// TIA Portal project "1215C_BREAKOUT_BOARD_IO-LINK_TOWERLIGHT" (V19) (continued)
REGION Network 6: Saving Selections
   RUNG wire#powerrail
      Contact( "DB005-HMI_Data".TowerLight.xSave_Config )
      wire#w1
      Move(in := #Seg2.iTempAnimation, out1 => "DB005-HMI_Data".TowerLight.Segment2.iSavedAnimate)
      Move(in := #Seg2.iTempSpeed, out1 => "DB003-IOLink_I/O".Outputs.TL_Byte_Array[13])
   END_RUNG
   RUNG wire#w1
      Move(in := #Seg2.iTempColour1, out1 => "DB003-IOLink_I/O".Outputs.TL_Byte_Array[15])
      Move(in := #Seg2.iTempColour2, out1 => "DB003-IOLink_I/O".Outputs.TL_Byte_Array[14])
      Move(in := #Seg2."iTempClrWidth%", out1 => "DB003-IOLink_I/O".Outputs.TL_Byte_Array[12])
   END_RUNG
   // the same network as SCL:
   IF "DB005-HMI_Data".TowerLight.xSave_Config THEN
       "DB005-HMI_Data".TowerLight.Segment2.iSavedAnimate := #Seg2.iTempAnimation;
       "DB003-IOLink_I/O".Outputs.TL_Byte_Array[13] := #Seg2.iTempSpeed;
       "DB003-IOLink_I/O".Outputs.TL_Byte_Array[15] := #Seg2.iTempColour1;
       "DB003-IOLink_I/O".Outputs.TL_Byte_Array[14] := #Seg2.iTempColour2;
       "DB003-IOLink_I/O".Outputs.TL_Byte_Array[12] := #Seg2."iTempClrWidth%";
   END_IF;
END_REGION

REGION Network 7: ================= SEGMENT_THREE =================
END_REGION

REGION Network 8: While making selections
   RUNG wire#powerrail
      { S7_Templates := "SrcType := UInt" } EQ_Contact(in1 := "DB005-HMI_Data".iScreen_Number, in2 := 9)
      wire#w1
      Move(in := "DB005-HMI_Data".TowerLight.Segment3.iAnimate, out1 => #Seg3.iTempAnimation)
      Move(in := "DB005-HMI_Data".TowerLight.Segment3.iSpeed, out1 => #Seg3.iTempSpeed)
   END_RUNG
   RUNG wire#w1
      Move(in := "DB005-HMI_Data".TowerLight.Segment3.iColour1, out1 => #Seg3.iTempColour1)
      Move(in := "DB005-HMI_Data".TowerLight.Segment3.iColour2, out1 => #Seg3.iTempColour2)
      Move(in := "DB005-HMI_Data".TowerLight.Segment3."iClrWidth%", out1 => #Seg3."iTempClrWidth%")
   END_RUNG
   // the same network as SCL:
   IF "DB005-HMI_Data".iScreen_Number = 9 THEN
       #Seg3.iTempAnimation := "DB005-HMI_Data".TowerLight.Segment3.iAnimate;
       #Seg3.iTempSpeed := "DB005-HMI_Data".TowerLight.Segment3.iSpeed;
       #Seg3.iTempColour1 := "DB005-HMI_Data".TowerLight.Segment3.iColour1;
       #Seg3.iTempColour2 := "DB005-HMI_Data".TowerLight.Segment3.iColour2;
       #Seg3."iTempClrWidth%" := "DB005-HMI_Data".TowerLight.Segment3."iClrWidth%";
   END_IF;
END_REGION

REGION Network 9: Saving Selections
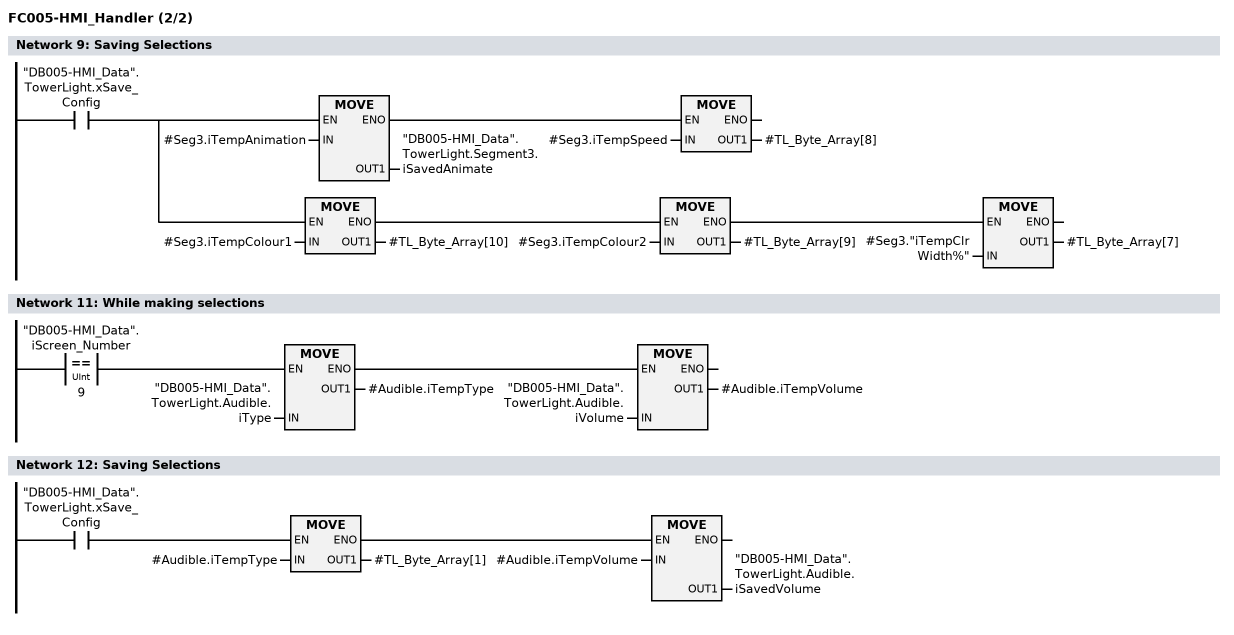
   RUNG wire#powerrail
      Contact( "DB005-HMI_Data".TowerLight.xSave_Config )
      wire#w1
      Move(in := #Seg3.iTempAnimation, out1 => "DB005-HMI_Data".TowerLight.Segment3.iSavedAnimate)
      Move(in := #Seg3.iTempSpeed, out1 => #TL_Byte_Array[8])
   END_RUNG
   RUNG wire#w1
      Move(in := #Seg3.iTempColour1, out1 => #TL_Byte_Array[10])
      Move(in := #Seg3.iTempColour2, out1 => #TL_Byte_Array[9])
      Move(in := #Seg3."iTempClrWidth%", out1 => #TL_Byte_Array[7])
   END_RUNG
   // the same network as SCL:
   IF "DB005-HMI_Data".TowerLight.xSave_Config THEN
       "DB005-HMI_Data".TowerLight.Segment3.iSavedAnimate := #Seg3.iTempAnimation;
       #TL_Byte_Array[8] := #Seg3.iTempSpeed;
       #TL_Byte_Array[10] := #Seg3.iTempColour1;
       #TL_Byte_Array[9] := #Seg3.iTempColour2;
       #TL_Byte_Array[7] := #Seg3."iTempClrWidth%";
   END_IF;
END_REGION

REGION Network 10: ================= AUDIBLE =================
END_REGION

REGION Network 11: While making selections
   RUNG wire#powerrail
      { S7_Templates := "SrcType := UInt" } EQ_Contact(in1 := "DB005-HMI_Data".iScreen_Number, in2 := 9)
      Move(in := "DB005-HMI_Data".TowerLight.Audible.iType, out1 => #Audible.iTempType)
      Move(in := "DB005-HMI_Data".TowerLight.Audible.iVolume, out1 => #Audible.iTempVolume)
   END_RUNG
   // the same network as SCL:
   IF "DB005-HMI_Data".iScreen_Number = 9 THEN
       #Audible.iTempType := "DB005-HMI_Data".TowerLight.Audible.iType;
       #Audible.iTempVolume := "DB005-HMI_Data".TowerLight.Audible.iVolume;
   END_IF;
END_REGION

REGION Network 12: Saving Selections
   RUNG wire#powerrail
      Contact( "DB005-HMI_Data".TowerLight.xSave_Config )
      Move(in := #Audible.iTempType, out1 => #TL_Byte_Array[1])
      Move(in := #Audible.iTempVolume, out1 => "DB005-HMI_Data".TowerLight.Audible.iSavedVolume)
   END_RUNG
   // the same network as SCL:
   IF "DB005-HMI_Data".TowerLight.xSave_Config THEN
       #TL_Byte_Array[1] := #Audible.iTempType;
       "DB005-HMI_Data".TowerLight.Audible.iSavedVolume := #Audible.iTempVolume;
   END_IF;
END_REGION
END_FUNCTION

// ===== library types =====

// folder: S7-1200/1500/Lib/S7-1200/1500/Common

FUNCTION_BLOCK "IO_LINK_DEVICE"   // FB50001, SCL
TITLE = IO_LINK_DEVICE
{ S7_Optimized_Access := 'TRUE' }
AUTHOR : SUP_FA
FAMILY : IO-Link
VERSION : 3.0
// Function block to read and write acyclic data on devices with IO-Link used on SIMATIC S7 controllers. (former IO_LINK_CALL)
   VAR_INPUT
      REQ : Bool;   // request function / Request Function / Neuer Auftrag
      ID : HW_IO;   // hardware identifier of IO-Link master module (HW_IO) from hw-config / Hardwarekennung des IOL-Master Moduls (HW_IO) aus HW-Konfiguration
      CAP : DInt := DINT#0;   // Client Access Point (CAP), for ET200 always 227 decimal / Client Access Point (CAP), bei ET200 immer 227 dez
      RD_WR : Bool;   // read and write access on IO-Link device 0: read, 1: write / Lese und Schreibzugriff auf IO-Link Device 0: Lesen, 1: schreiben
      PORT : Int := INT#0;   // number of port on IO-Link master module (ET200SP = 0..4) / Port/ Kanalnummer an dem das IO-Link Device betrieben wird. (ET200 = 0 .. 4)
      IOL_INDEX : Int := INT#0;   // address parameter Index (IO-Link Device) 0..32767 IOL-D, 65535 port functions / Adressparameter Index (IO-Link Device) 0..32767 IOL-D, 65535 port functions
      IOL_SUBINDEX : Int := INT#0;   // address parameter Subindex (IO-Link Device) 0 full record; 1-255 single parameter / Adressparameter Subindex (IO-Link Device) 0 ges. Record; 1-255 einz. Parameter
      LEN : Int := INT#0;   // length of writing data (netto data) / Länge der zu schreibenden Daten (Nettodaten)
   END_VAR
   VAR_OUTPUT
      DONE_VALID : Bool;   // validity 0: data invalid ; 1: data valid / Gültigkeit 0: Daten nicht gültig; 1: Daten gültig
      BUSY : Bool;   // 0: request finish 1: request in progress / 0: Auftrag abgeschlossen 1: Auftrag in Bearbeitung
      ERROR : Bool;   // Error Flag = 0: no error; 1: function aborted with error / Fehler Flag 0: kein Fehler; 1: Abbruch der Funktion mit Fehler
      STATUS : DWord := DW#16#00000000;   // DP/ PNIO - error status ; ERROR Flag = 1 - communication error status in detail / DP/ PNIO - Fehlerstatus; ERROR Flag = 1 - detaillierter Kommunikationsfehlerstatus
      IOL_STATUS : DWord := DW#16#00000000;   // IO-Link error status; ERROR flag = 1: IO-Link error status in detail / IO-Link Fehlerstatus; ERROR Flag = 1 - detaillierte IO-Link Fehlerstatus
      RD_LEN : Int := INT#0;   // length of read data record (number of bytes) / Länge des gelesenen Datensatzes (Anzahl Bytes)
   END_VAR
   VAR_IN_OUT
      RECORD_IOL_DATA : Array[0..231] of Byte;   // data area for reading / writing data (max. 232 byte) / Datenbereich für LESEN / SCHREIBEN (max. 232 Byte)
   END_VAR
   VAR
      RDREC_Function : RDREC;   // system function "read data record" (former SFB52) / Funktion Datensatz lesen (ehemals SFB52)
      WRREC_Function : WRREC;   // system function "write data record" (former SFB53) / Funktion Datensatz schreiben (ehemals SFB53)
      TP_poll : TP_TIME;   // poll rate read data record / Pollzeit für "Datensatz lesen"
      TON_monitoring : TON_TIME;   // request monitoring time / Überwachungszeit für Aufträge
      rdrec : Struct   // internal structure for RDREC / interne Struktur für RDREC
         valid : Bool;   // Function performed
         busy : Bool;   // Function busy
         error : Bool;   // Error flag
         status : DWord;   // Function result/error message
         length : UInt;   // Length of the fetched data record
      END_STRUCT;
      wrrec : Struct   // internal structure for WRREC / interne Struktur für WRREC
         length : UInt;   // length of write data record
         done : Bool;   // Function performed
         busy : Bool;   // Function busy
         error : Bool;   // Error flag
         status : DWord;   // Function result/error message
      END_STRUCT;
      read : Struct   // data area for reading data / Datenbereich für Lesedaten
         header : Struct
            CALL : Struct   // header for read/write data record
               Extended_Function_Num : Byte := 16#8;   // extended function number (fix coded 08h)
               Port : Byte;   // variable port (user interface) 0...255
               FI_Index : Word := 16#FE4A;   // FI index (fix coded 65098)
            END_STRUCT;
            IOL : Struct   // header for IO-Link
               Control : Byte;   // RD_WR = 0 = read = Control:=0x03 / / RD_WR = 1 = write = Control:=0x02
               Index_HighByte : Byte;   // index of data record 0…32767 (high byte)
               Index_LowByte : Byte;   // index of data record 0…32767 (low byte)
               Subindex : Byte;   // subindex for data record 0...255
            END_STRUCT;
         END_STRUCT;
         data : Array[0..231] of Byte;
      END_STRUCT;
      write : Struct   // data area for writing data / Datenbereich für Schreibdaten
         header : Struct
            CALL : Struct   // header for read/write data record
               Extended_Function_Num : Byte := 16#8;   // extended function number (fix coded 08h)
               Port : Byte;   // variable port (user interface) 0...255
               FI_Index : Word := 16#FE4A;   // FI index (fix coded 65098)
            END_STRUCT;
            IOL : Struct   // header for IO-Link
               Control : Byte;   // RD_WR = 0 = read = Control:=0x03 / / RD_WR = 1 = write = Control:=0x02
               Index_HighByte : Byte;   // index of data record 0…32767 (high byte)
               Index_LowByte : Byte;   // index of data record 0…32767 (low byte)
               Subindex : Byte;   // subindex for data record 0...255
            END_STRUCT;
         END_STRUCT;
         data : Array[0..231] of Byte;
      END_STRUCT;
      sequencecontrol : Int := INT#0;   // number of sequence control
      typeofrequest : Int := INT#0;   // type of request (0=Read, 1=Write)
      R_TRIG_REQ : Bool;   // impulse start new request / Impuls für neuen Auftrag starten
      R_TRIG_REQ_old : Bool;   // old value of REQ (previous cycle) / Flankenmerker
      F_TRIG_poll : Bool;   // impulse poll read data record (response) / Impuls für Pollen "Datensatz lesen"
      F_TRIG_poll_old : Bool;   // old value of Poll (previous cycle) / Flankenmerker
   END_VAR
   VAR_TEMP
      retval : Int;   // function return value / Variable für Rückgabewerte von Funktionen
      tmpWORD : Word;   // data type WORD for temporarily use / Datentyp WORD zur temporären Verwendung
      tmpDWORD : DWord;   // data type DWORD for temporarily use / Datentyp DWORD zur temporären Verwendung
      tmpINT : Int;   // data type INT for temporarily use / Datentyp INT zur temporären Verwendung
      i : Int;   // run tag for counting loops / Laufvariable für for-Schleifen
   END_VAR
BEGIN
   (*---------------------------------------------------------------------------------------------------------------------
   SIEMENS AG
   ©Copyright 2015. All Rights Reserved.
   -----------------------------------------------------------------------------------------------------------------------
   Limitation of liability
   This software was developed with largest care. However, the author can not guarantee, that the software runs under
   each version of STEP7 on each PLC flawlessly.
   There is no warranty for the software, to the extent permitted by applicable law. The copyright holder provides the
   software "as is" without warranty of any kind, either expressed or implied, including, but not limited to, the implied
   warranties of merchantability and fitness for a particular purpose. The entire risk as to the quality and performance
   of the software is with you. Should the software prove defective, you assume the cost of all necessary servicing,
   repair or correction. In no event unless required by applicable law will the copyright holder be liable to you for
   damages, including any general, special, incidental or consequential damages arising out of the use or inability to
   use the software (including but not limited to loss of data or data being rendered inaccurate or losses sustained by
   you or third parties or a failure of the software to operate with any other programs), even if such holder or other
   party has been advised of the possibility of such damages.
   Permission to use or copy this software for any purpose is hereby granted without fee, provided the above notices are
   retained on all copies. Permission to modify the code and to distribute modified code is granted, provided the above
   notices are retained, and a notice that the code was modified is included with the above copyright notice.
   -----------------------------------------------------------------------------------------------------------------------
   Functionality provided by this source (short description):
   Function block IO_LINK_DEVICE - used to read and write of acyclic data records on devices with IO-Link.
   Note:
   To read data records, the IO-Link master modules needs to know which data record is required. Therefore it is necessary
   to send at first a request via write data record (only header of 8 byte). As response the IO-Link master module
   will send the required data record.

   Status:     Released (tested)
   File name:  IO_LINK_DEVICE
   System :    SIMATIC S7-1200/1500
   Version :   3.0
   -----------------------------------------------------------------------------------------------------------------------
   Script to be stored on level ... in project (mark appropriate levels with [x] below)
   [ ] External
   [ ] All levels possible
   [x] Project level
   [ ] Controller level
   [ ] Device level
   [ ] Subobject level
   -----------------------------------------------------------------------------------------------------------------------
   Restrictions, known limitations:
   The limitation of 240 byte is based on PROFIBUS DP protocol. With PROFINET IO there wouldn't no limit but because of 
   compatibility reason it wasn't changed.
     - header =   8 byte
     - data   = 232 byte
   -----------------------------------------------------------------------------------------------------------------------
   Requirements, prerequisites, External resources used: nothing
   -----------------------------------------------------------------------------------------------------------------------
   Change log table (latest change is at the bottom OF the list):
   Version Date Changes applied
   V2.0.0 <2013-09-30> First created with TIA Portal V12 SP1
   V2.1.0 <2014-03-14> Upgrade system function 'WRREC' from V1.0 to V1.1 and released for TIA Portal V13
   V3.0.0 <2015-02-28> Upgrade and released for TIA Portal V13 SP1 (without backup/restore master parameter)
   V3.0.2 <2015-07-07> Change of #IOL_INDEX and #Port lower boundry to 0
   ---------------------------------------------------------------------------------------------------------------------*)

   (*---------------------------------------------------------------------------------------------------------------------
   Description of programmed IO-Link error codes
   8000 = time out
   8001 = wrong port
   8002 = wrong index
   8003 = wrong subindex
   8005 = wrong length for write data record
   8006 = wrong length for read data record
   8052 = error during reading data record
   8053 = error during writing data record
   All other codes are coming from a higher level!
   ---------------------------------------------------------------------------------------------------------------------*)

   (*---------------------------------------------------------------------------------------------------------------------
               NEW REQUEST
   ---------------------------------------------------------------------------------------------------------------------*)
   // detection rising edge of "REQ"
   #R_TRIG_REQ := #REQ = TRUE AND #R_TRIG_REQ_old = FALSE;
   #R_TRIG_REQ_old := #REQ = TRUE;

   // start new request if not busy
   IF #R_TRIG_REQ = TRUE AND #sequencecontrol = 0 THEN
       // Freeze record ID and CAP
       #WRREC_Function.ID := #ID;
       #WRREC_Function.INDEX := #CAP;
       #RDREC_Function.ID := #ID;
       #RDREC_Function.INDEX := #CAP;

       // Initialize outputs
       #DONE_VALID := FALSE;
       #BUSY := TRUE;
       #ERROR := FALSE;
       #STATUS := DW#16#00000000;
       #IOL_STATUS := DW#16#00000000;
       #RD_LEN := INT#0;

       // Initialize data area
       #read.header.CALL.Port := B#16#0;
       #read.header.IOL.Index_LowByte := B#16#0;
       #read.header.IOL.Index_HighByte := B#16#0;
       #read.header.IOL.Subindex := B#16#0;
       #i := INT#0; // initialize loop counter      
       FOR #i := 0 TO 231 DO
           #write.data[#i] := B#16#0;
           #read.data[#i] := B#16#0;
       END_FOR;

   (*---------------------------------------------------------------------------------------------------------------------
       Setup IO-LINK Call needs a specific header
   ---------------------------------------------------------------------------------------------------------------------*)
   // setup CALL header
   #write.header.CALL.Extended_Function_Num := 16#08;  // extended function number (fix coded 08h)
   #write.header.CALL.Port := INT_TO_BYTE(#PORT);  // 1..63 = PORT number, 64..255=reserved
   #write.header.CALL.FI_Index := 65098;  // IOL-Header is following (fix coded 65098)

   // setup IOL header 
   // CONTROL = please see below at BODY
   // INDEX
   #write.header.IOL.Index_LowByte := INT_TO_BYTE(#IOL_INDEX);
   #tmpWORD := INT_TO_WORD(#IOL_INDEX);
   #tmpWORD := SHR(IN := #tmpWORD, N := 8);
   #write.header.IOL.Index_HighByte := WORD_TO_BYTE(#tmpWORD);
   // SUBINDEX
   #write.header.IOL.Subindex := INT_TO_BYTE(#IOL_SUBINDEX);

   // BODY (data max. 232 Byte, Array 0..231 of Byte) 
   IF #RD_WR = TRUE THEN
       // IO-Link write data record requested, copy data from "RECORD_IOL_DATA"
       #write.header.IOL.Control := B#16#02; // CONTROL B#16#02 = write data record
       #wrrec.length := INT_TO_UINT(#LEN) + UINT#8;  // data length header + data = IO-Link write data record
       #typeofrequest := 2; // write data record
       // copy IOL_RECORD_DATA in working area
       #i := INT#0;    // initialize loop counter 
       FOR #i := 0 TO #LEN - 1 DO
           #write.data[#i] := #RECORD_IOL_DATA[#i];
       END_FOR;
   ELSE
       // IO-Link read data record requested
       #write.header.IOL.Control := 16#03;  // CONTROL 16#03 = read data record
       #wrrec.length := UINT#8; // data length only header = IO-Link read data record
       #typeofrequest := 1; // read data record        
   END_IF;
   #sequencecontrol := 1;  // Start sequence
   ELSE
       ;
   END_IF;

   (*---------------------------------------------------------------------------------------------------------------------
               SEQUENCE CONTROL
   ---------------------------------------------------------------------------------------------------------------------*)
   CASE #sequencecontrol OF
       1:  // Check input parameter        
           IF #PORT < INT#0 OR #PORT > INT#63 THEN // PORT (Wrong port address = 0x8001)
               #ERROR := TRUE;
               #IOL_STATUS := DW#16#80010000;
               #sequencecontrol := 99; // aborting function with error
           ELSIF #IOL_INDEX < INT#0 OR #IOL_INDEX > INT#32767 THEN    // INDEX (Wrong index = 0x8002)
               #ERROR := TRUE;
               #IOL_STATUS := DW#16#80020000;
               #sequencecontrol := 99; // aborting function with error
           ELSIF #IOL_SUBINDEX < INT#0 OR #IOL_SUBINDEX > INT#255 THEN    // SUBINDEX (Wrong subindex = 0x8003)
               #ERROR := TRUE;
               #IOL_STATUS := DW#16#80030000;
               #sequencecontrol := 99; // aborting function with error
           ELSIF #typeofrequest = 2 AND (#LEN < 1 OR #LEN > 232) THEN  // LEN (wrong length for write data record = 0x8004)
               #ERROR := TRUE;
               #IOL_STATUS := DW#16#80050000;
               #sequencecontrol := 99; // aborting function with error
           ELSIF #typeofrequest = 1 AND (#LEN < 0 OR #LEN > 232) THEN  // LEN (wrong length for read data record = 0x8005)
               #ERROR := TRUE;
               #IOL_STATUS := DW#16#80060000;
               #sequencecontrol := 99; // aborting function with error
           ELSE    // all input parameter are right
               #sequencecontrol := 2;
           END_IF;

       2:  (*-------------------------------------------------------------------------------------------------------------
           WRREC = Write Data Record
           Note:
           To read data records, the IO-Link master modules needs to know which PORT is required. Therefore it is necessary
           to send at first a request via write data record (header, 8 byte). As response the IO-Link master module will 
           send the required data record.
           -------------------------------------------------------------------------------------------------------------*)
           #WRREC_Function(REQ := TRUE,
                           LEN := #wrrec.length,
                           DONE => #wrrec.done,
                           BUSY => #wrrec.busy,
                           ERROR => #wrrec.error,
                           STATUS => #wrrec.status,
                           RECORD := #write);
           // output status during write data record
           IF #wrrec.busy THEN
               #STATUS := #wrrec.status;
               #IOL_STATUS := DW#16#00020000;  // 0002 = writing in progress 
           ELSIF #wrrec.error THEN
               #tmpDWORD := #wrrec.status AND DW#16#00FFFF00;  // filter status
               IF #tmpDWORD = DW#16#0080C200 THEN    // if resource #BUSY (#STATUS=80C2), then ... 
                   #sequencecontrol := 3;  // ... repeat write data record
               ELSE
                   #ERROR := TRUE;
                   #STATUS := #wrrec.status;   // ... otherwise output error status of "WRREC"
                   #IOL_STATUS := DW#16#80530000;  // ... with note '8053' = error status of "WRREC"
                   #sequencecontrol := 99; // aborting function with error
               END_IF;
           ELSIF #wrrec.done = TRUE THEN   // wait for write data record finish without error
               #TP_poll(IN := TRUE,
                        PT := T#100ms);    // poll for response
               #sequencecontrol := 4;
           ELSE
               ;
           END_IF;

       3:  // repeat write data record because resource was busy
           #WRREC_Function(REQ := FALSE);
           #sequencecontrol := 2;

       4:  // wait and poll for response = Read Data Record (RDREC)
           #WRREC_Function(REQ := FALSE);
           #TP_poll(IN := TRUE,
                    PT := T#100ms);

           // if poll rate executed then start read data record (on falling edge)
           #F_TRIG_poll := #TP_poll.Q = FALSE AND #F_TRIG_poll_old = TRUE;
           #F_TRIG_poll_old := #TP_poll.Q = TRUE;

           // RDREC = Read Data Record
           #RDREC_Function(REQ := #F_TRIG_poll,
                           MLEN := UINT#0, // length = 0 = read all data which are available
                           VALID => #rdrec.valid,
                           BUSY => #rdrec.busy,
                           ERROR => #rdrec.error,
                           STATUS => #rdrec.status,
                           LEN => #rdrec.length,
                           RECORD := #read);
           // output status during read data record
           IF #rdrec.busy THEN
               #STATUS := #rdrec.status;
               #IOL_STATUS := DW#16#00030000; // 16#0003 = reading in progress
           ELSIF #rdrec.error = TRUE THEN
               #tmpDWORD := #rdrec.status AND DW#16#00FFFF00;  // filter status
               IF #tmpDWORD = DW#16#0080C200 THEN  // if resource busy (status=80C2), then ... 
                   #sequencecontrol := 5;  // ... repeat read data record / continue polling
               ELSE
                   #ERROR := TRUE;
                   #STATUS := #rdrec.status;   // ... otherwise output error code of "RDREC"
                   #IOL_STATUS := DW#16#80520000;  // ... with note '8052' = error status of "RDREC"
                   #sequencecontrol := 99; // aborting function with error
               END_IF;
           ELSIF #rdrec.valid THEN
               IF  // check the response wether it matches the request (compare PORT, INDEX and SUBINDEX)
                   (#write.header.CALL.Port <> #read.header.CALL.Port) OR
                   (#write.header.IOL.Index_HighByte <> #read.header.IOL.Index_HighByte) OR
                   (#write.header.IOL.Index_LowByte <> #read.header.IOL.Index_LowByte) OR
                   (#write.header.IOL.Subindex <> #read.header.IOL.Subindex)
               THEN    // read data record don't match the request
                   #ERROR := TRUE;
                   #STATUS := #rdrec.status;
                   #IOL_STATUS := DW#16#70000000;  // output status '7000', no consistent data
                   #sequencecontrol := 99; // aborting function with error
               ELSIF #read.header.IOL.Control = B#16#80 THEN   // check the response for IO-Link errors
                   // State 0x80 = IOL_CALL_RES PDU shows IO-Link error detect
                   #ERROR := TRUE;
                   #STATUS := DW#16#00000000;
                   #IOL_STATUS.%B3 := #read.data[0];   // IO-Link master error code
                   #IOL_STATUS.%B2 := #read.data[1];   // IO-Link master error code
                   #IOL_STATUS.%B1 := #read.data[2];  // IO-Link device error code
                   #IOL_STATUS.%B0 := #read.data[3];  // IO-Link device additional error code

                   #sequencecontrol := 99; // aborting function with error
               ELSE    // read data are valid = output
                   #DONE_VALID := TRUE;
                   #BUSY := FALSE;
                   #ERROR := FALSE;
                   #STATUS := DW#16#00000000;
                   #IOL_STATUS := DW#16#00000000;  // request finished

                   IF #typeofrequest = 1 THEN
                       #RD_LEN := UINT_TO_INT(#rdrec.length - UINT#8);  // device parameter cover header and data,
                       // only data will be output
                       #i := INT#0; // initialize loop counter
                       FOR #i := 0 TO UINT_TO_INT(#rdrec.length - UINT#8 - UINT#1) DO
                           #RECORD_IOL_DATA[#i] := #read.data[#i];
                       END_FOR;
                   ELSE
                       ;
                   END_IF;
                   #sequencecontrol := 98;
               END_IF;
           ELSE
               ;
           END_IF;

       5:  // poll again for response because resource was busy
           #TP_poll(IN := FALSE,
                    PT := T#100ms);
           #RDREC_Function(REQ := FALSE,
                           RECORD := #read);
           #sequencecontrol := 4;  // ... repeat read data record / continue polling   

       98: // request done successfully
           #TP_poll(IN := FALSE,
                    PT := T#100ms);
           #RDREC_Function(REQ := FALSE,
                           RECORD := #read);
           IF #REQ = FALSE THEN
               #DONE_VALID := FALSE;
               #BUSY := FALSE;
               #ERROR := FALSE;
               #RD_LEN := INT#0;
               #STATUS := DW#16#00000000;
               #IOL_STATUS := DW#16#00010000; // ready for new request
               #sequencecontrol := 0;
               #typeofrequest := 0;
           ELSE
               ;
           END_IF;

       99: // Function aborted with error
           #TP_poll(IN := FALSE,
                    PT := T#100ms);
           #WRREC_Function(REQ := FALSE);
           #RDREC_Function(REQ := FALSE,
                           RECORD := #read);
           #DONE_VALID := FALSE;
           #BUSY := FALSE;
           #RD_LEN := INT#0;
           #sequencecontrol := 0;
           #typeofrequest := 0;

       ELSE  // no relevant case, ready for new request
           #WRREC_Function(REQ := FALSE);
           #RDREC_Function(REQ := FALSE,
                           RECORD := #read);
           #TP_poll(IN := FALSE,
                    PT := T#100ms);
           #TON_monitoring(IN := FALSE,
                           PT := T#20s);
           #sequencecontrol := 0;
           #typeofrequest := 0;
   END_CASE;

   (*---------------------------------------------------------------------------------------------------------------------
               MONITORING
   ---------------------------------------------------------------------------------------------------------------------*)
   #TON_monitoring(IN := #sequencecontrol > 0 AND #sequencecontrol < 98,
                   PT := T#20s);
   IF #TON_monitoring.Q THEN
       #ERROR := TRUE;
       #IOL_STATUS := DW#16#80000000; // request time out       
       #sequencecontrol := 99; // aborting function with error
   END_IF;
END_FUNCTION_BLOCK

(* ===== HMI "HMI_RT_1" =====
system functions are stored by id; their names below are inferred from use
connection "HMI_Connection": ETHERNET, SMART_S7_1200_OMS

HMI tags "PLC_Inputs"
   "DB001-PLC_I/O_Inputs_xDI0.0" : Bool = PLC "DB001-PLC_I/O".Inputs."xDI0.0", 100 ms
   "DB001-PLC_I/O_Inputs_xDI0.1" : Bool = PLC "DB001-PLC_I/O".Inputs."xDI0.1", 100 ms
   "DB001-PLC_I/O_Inputs_xDI0.2" : Bool = PLC "DB001-PLC_I/O".Inputs."xDI0.2", 100 ms
   "DB001-PLC_I/O_Inputs_xDI0.3" : Bool = PLC "DB001-PLC_I/O".Inputs."xDI0.3", 100 ms
   "DB001-PLC_I/O_Inputs_xDI0.4" : Bool = PLC "DB001-PLC_I/O".Inputs."xDI0.4", 100 ms
   "DB001-PLC_I/O_Inputs_xDI0.5" : Bool = PLC "DB001-PLC_I/O".Inputs."xDI0.5", 100 ms
   "DB001-PLC_I/O_Inputs_xDI0.6" : Bool = PLC "DB001-PLC_I/O".Inputs."xDI0.6", 100 ms
   "DB001-PLC_I/O_Inputs_xDI0.7" : Bool = PLC "DB001-PLC_I/O".Inputs."xDI0.7", 100 ms
   "DB001-PLC_I/O_Inputs_xDI1.0" : Bool = PLC "DB001-PLC_I/O".Inputs."xDI1.0", 100 ms
   "DB001-PLC_I/O_Inputs_xDI1.1" : Bool = PLC "DB001-PLC_I/O".Inputs."xDI1.1", 100 ms
   "DB001-PLC_I/O_Inputs_xDI1.2" : Bool = PLC "DB001-PLC_I/O".Inputs."xDI1.2", 100 ms
   "DB001-PLC_I/O_Inputs_xDI1.3" : Bool = PLC "DB001-PLC_I/O".Inputs."xDI1.3", 100 ms
   "DB001-PLC_I/O_Inputs_xDI1.4" : Bool = PLC "DB001-PLC_I/O".Inputs."xDI1.4", 100 ms
   "DB001-PLC_I/O_Inputs_xDI1.5" : Bool = PLC "DB001-PLC_I/O".Inputs."xDI1.5", 100 ms

HMI tags "PLC_Outputs"
   "DB001-PLC_I/O_Outputs_xDQ0.0" : Bool = PLC "DB001-PLC_I/O".Outputs."xDQ0.0", 100 ms
   "DB001-PLC_I/O_Outputs_xDQ0.1" : Bool = PLC "DB001-PLC_I/O".Outputs."xDQ0.1", 100 ms
   "DB001-PLC_I/O_Outputs_xDQ0.2" : Bool = PLC "DB001-PLC_I/O".Outputs."xDQ0.2", 100 ms
   "DB001-PLC_I/O_Outputs_xDQ0.3" : Bool = PLC "DB001-PLC_I/O".Outputs."xDQ0.3", 100 ms
   "DB001-PLC_I/O_Outputs_xDQ0.4" : Bool = PLC "DB001-PLC_I/O".Outputs."xDQ0.4", 100 ms
   "DB001-PLC_I/O_Outputs_xDQ0.5" : Bool = PLC "DB001-PLC_I/O".Outputs."xDQ0.5", 100 ms
   "DB001-PLC_I/O_Outputs_xDQ0.6" : Bool = PLC "DB001-PLC_I/O".Outputs."xDQ0.6", 100 ms
   "DB001-PLC_I/O_Outputs_xDQ0.7" : Bool = PLC "DB001-PLC_I/O".Outputs."xDQ0.7", 100 ms
   "DB001-PLC_I/O_Outputs_xDQ1.0" : Bool = PLC "DB001-PLC_I/O".Outputs."xDQ1.0", 100 ms
   "DB001-PLC_I/O_Outputs_xDQ1.1" : Bool = PLC "DB001-PLC_I/O".Outputs."xDQ1.1", 100 ms

HMI tags "PLC_Analog"
   "AI0.0" : Word = PLC "AI0.0" AT %IW64, 100 ms
   "AQ0.0" : Word = PLC "AQ0.0" AT %QW64, 100 ms
   "DB001-PLC_I/O_Outputs_rAQ0.0_Scaled" : Real = PLC "DB001-PLC_I/O".Outputs."rAQ0.0_Scaled", 100 ms
   "DB001-PLC_I/O_Outputs_rAQ0.1_Scaled" : Real = PLC "DB001-PLC_I/O".Outputs."rAQ0.1_Scaled", 100 ms
   "AI0.1" : Word = PLC "AI0.1" AT %IW66, 100 ms
   "AQ0.1" : Word = PLC "AQ0.1" AT %QW66, 100 ms
   "DB001-PLC_I/O_Inputs_rAI0.0_Scaled" : Real = PLC "DB001-PLC_I/O".Inputs."rAI0.0_Scaled", 100 ms
   "DB001-PLC_I/O_Inputs_rAI0.1_Scaled" : Real = PLC "DB001-PLC_I/O".Inputs."rAI0.1_Scaled", 100 ms

HMI tags "PLC_DateTime"
   "DB002-DateTime_sCustomDate_DDMMYY" : String[254] = PLC "DB002-DateTime".sCustomDate_DDMMYY, 100 ms
   "DB002-DateTime_sCustomTime_HHMM" : String[254] = PLC "DB002-DateTime".sCustomTime_HHMM, 100 ms

HMI tags "HMI_Data"
   "DB005-HMI_Data_TowerLight_Audible_iType" : Int = PLC "DB005-HMI_Data".TowerLight.Audible.iType, 100 ms
   "DB005-HMI_Data_TowerLight_Audible_iVolume" : Int = PLC "DB005-HMI_Data".TowerLight.Audible.iVolume, 100 ms
   "DB005-HMI_Data_TowerLight_Segment1_iAnimate" : Int = PLC "DB005-HMI_Data".TowerLight.Segment1.iAnimate, 100 ms
   "DB005-HMI_Data_TowerLight_Segment1_iClrWidth%" : Int = PLC "DB005-HMI_Data".TowerLight.Segment1.iClrWidth%, 100 ms
   "DB005-HMI_Data_TowerLight_Segment1_iColour1" : Int = PLC "DB005-HMI_Data".TowerLight.Segment1.iColour1, 100 ms
   "DB005-HMI_Data_TowerLight_Segment1_iColour2" : Int = PLC "DB005-HMI_Data".TowerLight.Segment1.iColour2, 100 ms
   "DB005-HMI_Data_TowerLight_Segment1_iSpeed" : Int = PLC "DB005-HMI_Data".TowerLight.Segment1.iSpeed, 100 ms
   "DB005-HMI_Data_TowerLight_Segment2_iAnimate" : Int = PLC "DB005-HMI_Data".TowerLight.Segment2.iAnimate, 100 ms
   "DB005-HMI_Data_TowerLight_Segment2_iClrWidth%" : Int = PLC "DB005-HMI_Data".TowerLight.Segment2.iClrWidth%, 100 ms
   "DB005-HMI_Data_TowerLight_Segment2_iColour1" : Int = PLC "DB005-HMI_Data".TowerLight.Segment2.iColour1, 100 ms
   "DB005-HMI_Data_TowerLight_Segment2_iColour2" : Int = PLC "DB005-HMI_Data".TowerLight.Segment2.iColour2, 100 ms
   "DB005-HMI_Data_TowerLight_Segment2_iSpeed" : Int = PLC "DB005-HMI_Data".TowerLight.Segment2.iSpeed, 100 ms
   "DB005-HMI_Data_TowerLight_Segment3_iAnimate" : Int = PLC "DB005-HMI_Data".TowerLight.Segment3.iAnimate, 100 ms
   "DB005-HMI_Data_TowerLight_Segment3_iClrWidth%" : Int = PLC "DB005-HMI_Data".TowerLight.Segment3.iClrWidth%, 100 ms
   "DB005-HMI_Data_TowerLight_Segment3_iColour1" : Int = PLC "DB005-HMI_Data".TowerLight.Segment3.iColour1, 100 ms
   "DB005-HMI_Data_TowerLight_Segment3_iColour2" : Int = PLC "DB005-HMI_Data".TowerLight.Segment3.iColour2, 100 ms
   "DB005-HMI_Data_TowerLight_Segment3_iSpeed" : Int = PLC "DB005-HMI_Data".TowerLight.Segment3.iSpeed, 100 ms
   "DB005-HMI_Data_TowerLight_xSave_Config" : Bool = PLC "DB005-HMI_Data".TowerLight.xSave_Config, 100 ms
   "DB005-HMI_Data_iScreen_Number" : UInt = PLC "DB005-HMI_Data".iScreen_Number AT %DB1.DBW0, 100 ms

text list "ON/OFF": 0 'OFF'; 1 'ON'

text list "Animate": 0 'Off'; 1 'Steady'; 2 'Flash'; 3 '2Colour Flash'; 4 '2Colour Shift'; 5 'Ends Steady'; 6 'Ends Flash'; 7 'Scroll'; 8 'Center Scroll'; 9 'Bounce'; 10 'Center Bounce'; 11 'Intensity Sweep'; 12 '2Colour Sweep'; 13 'Spectrum'; 14 'Level Steady'; 15 'Level Flash'

text list "Colour1": 0 'Green'; 1 'Red'; 2 'Orange'; 3 'Amber'; 4 'Yellow'; 5 'Lime Green'; 6 'Spring Green'; 7 'Cyan'; 8 'Sky Blue'; 9 'Blue'; 10 'Violet'; 11 'Magenta'; 12 'Rose'; 13 'Daylight White'

text list "Colour2": 0 'Green'; 1 'Red'; 2 'Orange'; 3 'Amber'; 4 'Yellow'; 5 'Lime Green'; 6 'Spring Green'; 7 'Cyan'; 8 'Sky Blue'; 9 'Blue'; 10 'Violet'; 11 'Magenta'; 12 'Rose'; 13 'Daylight White'

text list "Speed": 0 'Medium'; 1 'Fast'; 2 'Slow'

text list "Type": 0 'Pulse'; 1 'Wobble'; 2 'Strobe'; 4 'Whoop'; 5 'Staccato'; 6 'Siren'; 8 'Continuous1'; 9 'Continuous2'; 16 'Jingle'; 17 'Melody1'; 18 'Melody2'; 19 'Melody3'

text list "Volume": 0 'Off'; 1 'Low'; 2 'Medium'; 3 'High'

screen "01-Home" 480x272, template "Main_Template"
   on GenerateScreen: SetTag("DB005-HMI_Data_iScreen_Number", 1)
   TextField "TextField_ProjectName" at 109,47 size 259x30; Text 'PLC BREAKOUT BOARD'
   TextField "Text field_DeviceInfo" at 21,85 size 435x52; Text '1215C DC/DC/DC -- 6ES7215-1AG40-0XB0 -- IP: 192.168.0.175/24 KTP400 HMI -- 6AV2123-2DB03-0AX0 -- IP: 192.168.0.176/24 IFM IO-LINK MASTER -- AL1100 -- IP: 192.168.0.177/24'
   TextField "Text field_Description" at 62,143 size 369x68; Text '- Displays the Digital & Analog I/O states, - Toggle Digital Outputs via HMI buttons, - Simulation of Analog Outputs via 20 step incriments, - Configuration & Control of IO-Link Tower Light via HMI.'
   Button "Button_ExitRuntime" at 384,227 size 92x40; TextOff 'EXIT RUNTIME'
      on Press: StopRuntime(0)

screen "02-Inputs1" 480x272, template "Main_Template"
   on GenerateScreen: SetTag("DB005-HMI_Data_iScreen_Number", 2)
   TextField "TextField_ScreenName" at 85,46 size 309x30; Text 'PLC DIGITAL INPUTS - 1of3'
   TextField "TextField_BankLetter" at 412,50 size 64x23; Text 'BANK A'
   Button "Button_Next" at 384,227 size 92x40; TextOff 'NEXT'
      on Press: ActivateScreen("03-Inputs2", 0)
   Group "Group_DI0.0" at 41,81 size 62x63
   Group "Group_DI0.1" at 153,81 size 62x63
   Group "Group_DI0.2" at 265,81 size 62x63
   Group "Group_DI0.3" at 377,81 size 62x63
   Group "Group_DI0.4" at 41,152 size 62x64
   Group "Group_DI0.5" at 153,152 size 62x64
   Group "Group_DI0.6" at 265,154 size 62x64
   Group "Group_DI0.7" at 377,154 size 62x64
   TextField "Text field_DI0.0" at 51,81 size 42x19; Text 'DI 0.0'
   Circle "Circle_DI0.0" at 54,103 size 36x36
      Appearance <- "DB001-PLC_I/O_Inputs_xDI0.0"
   TextField "Text field_DI0.1" at 163,81 size 42x19; Text 'DI 0.1'
   Circle "Circle_DI0.1" at 166,103 size 36x36
      Appearance <- "DB001-PLC_I/O_Inputs_xDI0.1"
   TextField "Text field_DI0.2" at 275,81 size 42x19; Text 'DI 0.2'
   Circle "Circle_DI0.2" at 278,103 size 36x36
      Appearance <- "DB001-PLC_I/O_Inputs_xDI0.2"
   TextField "Text field_DI0.3" at 387,81 size 42x19; Text 'DI 0.3'
   Circle "Circle_DI0.3" at 390,103 size 36x36
      Appearance <- "DB001-PLC_I/O_Inputs_xDI0.3"
   TextField "Text field_DI0.4" at 51,152 size 42x19; Text 'DI 0.4'
   Circle "Circle_DI0.4" at 54,174 size 36x36
      Appearance <- "DB001-PLC_I/O_Inputs_xDI0.4"
   TextField "Text field_DI0.5" at 163,152 size 42x19; Text 'DI 0.5'
   Circle "Circle_DI0.5" at 166,174 size 36x36
      Appearance <- "DB001-PLC_I/O_Inputs_xDI0.5"
   TextField "Text field_DI0.6" at 275,154 size 42x19; Text 'DI 0.6'
   Circle "Circle_DI0.6" at 278,176 size 36x36
      Appearance <- "DB001-PLC_I/O_Inputs_xDI0.6"
   TextField "Text field_DI0.7" at 387,154 size 42x19; Text 'DI 0.7'
   Circle "Circle_DI0.7" at 390,176 size 36x36
      Appearance <- "DB001-PLC_I/O_Inputs_xDI0.7"

